// TIA Portal project "Factory_Project_V17" (V17) (continued)
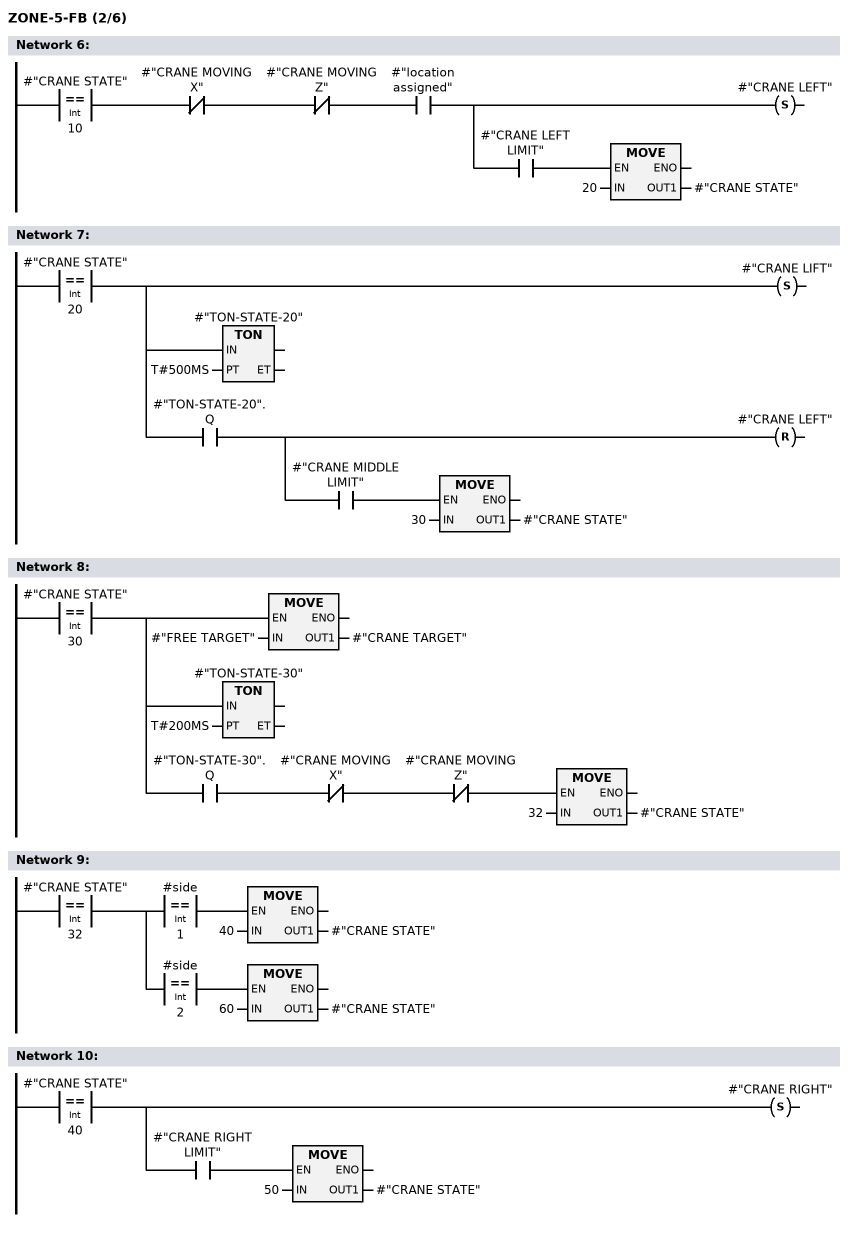
   RUNG wire#powerrail
      { S7_Templates := "SrcType := Int" } EQ_Contact(in1 := #"CRANE STATE", in2 := 10)
      I_Contact( #"CRANE MOVING X" )
      I_Contact( #"CRANE MOVING Z" )
      Contact( #"location assigned" )
      wire#w1
      S_Coil( #"CRANE LEFT" )
   END_RUNG
   RUNG wire#w1
      Contact( #"CRANE LEFT LIMIT" )
      Move(in := 20, out1 => #"CRANE STATE")
   END_RUNG
   // the same network as SCL:
   #_w1 := (#"CRANE STATE" = 10) AND NOT #"CRANE MOVING X" AND NOT #"CRANE MOVING Z" AND #"location assigned";
   IF #_w1 THEN #"CRANE LEFT" := TRUE; END_IF;
   IF #_w1 AND #"CRANE LEFT LIMIT" THEN #"CRANE STATE" := 20; END_IF;
END_REGION

REGION Network 7
   #_w1 := #"CRANE STATE" = 20;
   IF #_w1 THEN #"CRANE LIFT" := TRUE; END_IF;
   #"TON-STATE-20"(IN := #_w1, PT := T#500MS);   // TON
   #_w2 := #_w1 AND #"TON-STATE-20".Q;
   IF #_w2 THEN #"CRANE LEFT" := FALSE; END_IF;
   IF #_w2 AND #"CRANE MIDDLE LIMIT" THEN #"CRANE STATE" := 30; END_IF;
END_REGION

REGION Network 8
   #_w1 := #"CRANE STATE" = 30;
   IF #_w1 THEN #"CRANE TARGET" := #"FREE TARGET"; END_IF;
   #"TON-STATE-30"(IN := #_w1, PT := T#200MS);   // TON
   IF #_w1 AND #"TON-STATE-30".Q AND NOT #"CRANE MOVING X" AND NOT #"CRANE MOVING Z" THEN
       #"CRANE STATE" := 32;
   END_IF;
END_REGION

REGION Network 9
   RUNG wire#powerrail
      { S7_Templates := "SrcType := Int" } EQ_Contact(in1 := #"CRANE STATE", in2 := 32)
      wire#w1
      { S7_Templates := "SrcType := Int" } EQ_Contact(in1 := #side, in2 := 1)
      Move(in := 40, out1 => #"CRANE STATE")
   END_RUNG
   RUNG wire#w1
      { S7_Templates := "SrcType := Int" } EQ_Contact(in1 := #side, in2 := 2)
      Move(in := 60, out1 => #"CRANE STATE")
   END_RUNG
   // the same network as SCL:
   #_w1 := #"CRANE STATE" = 32;
   IF #_w1 AND (#side = 1) THEN #"CRANE STATE" := 40; END_IF;
   IF #_w1 AND (#side = 2) THEN #"CRANE STATE" := 60; END_IF;
END_REGION

REGION Network 10
   RUNG wire#powerrail
      { S7_Templates := "SrcType := Int" } EQ_Contact(in1 := #"CRANE STATE", in2 := 40)
      wire#w1
      S_Coil( #"CRANE RIGHT" )
   END_RUNG
   RUNG wire#w1
      Contact( #"CRANE RIGHT LIMIT" )
      Move(in := 50, out1 => #"CRANE STATE")
   END_RUNG
   // the same network as SCL:
   #_w1 := #"CRANE STATE" = 40;
   IF #_w1 THEN #"CRANE RIGHT" := TRUE; END_IF;
   IF #_w1 AND #"CRANE RIGHT LIMIT" THEN #"CRANE STATE" := 50; END_IF;
END_REGION

REGION Network 11
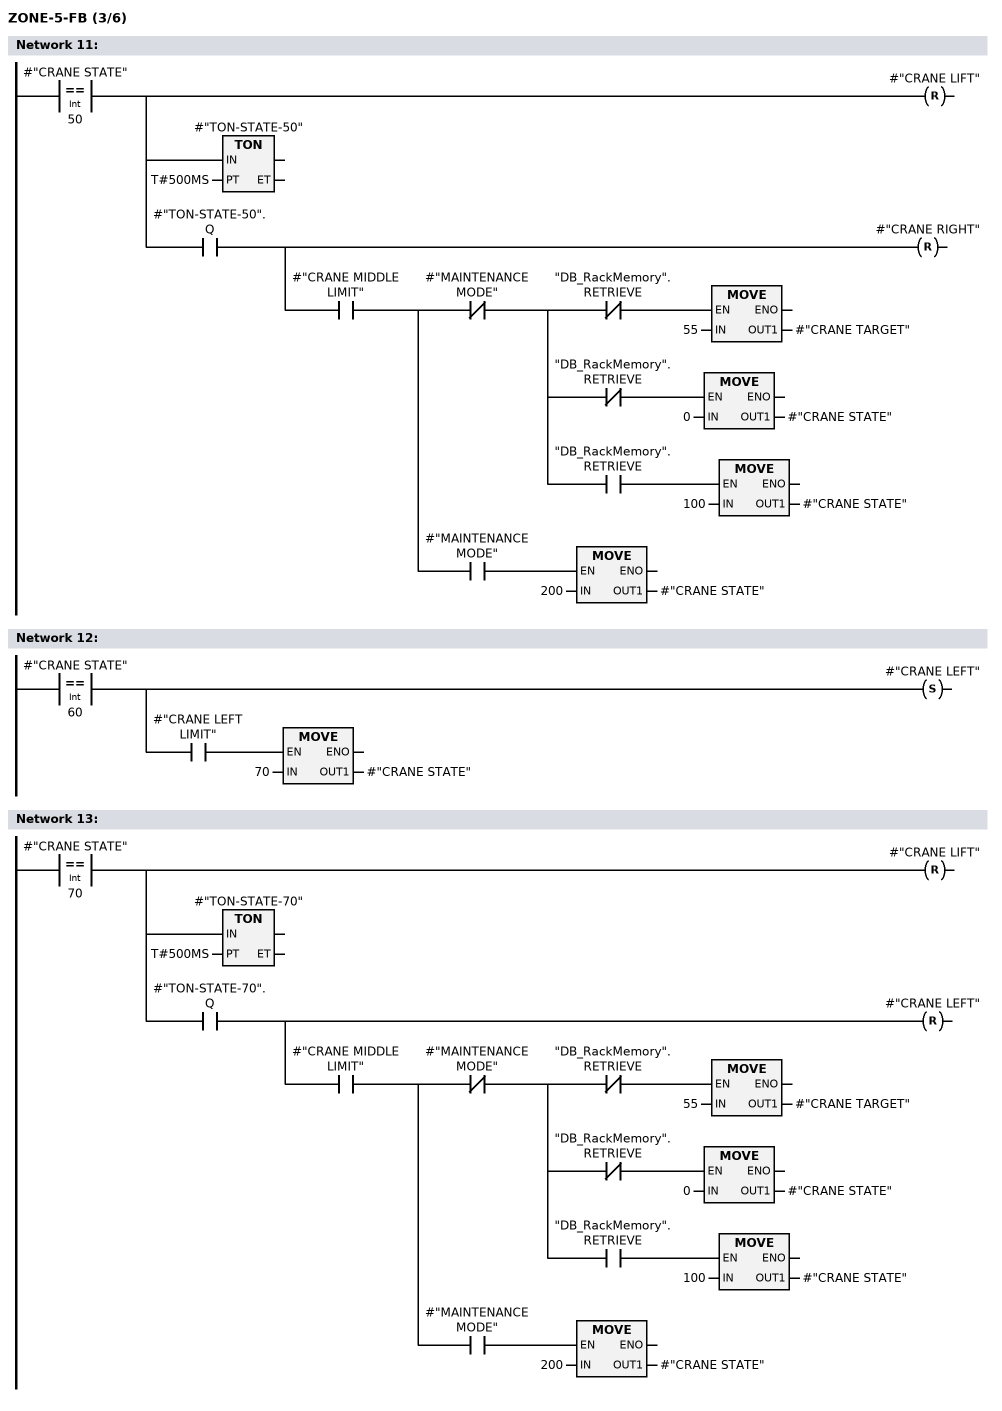
   #_w1 := #"CRANE STATE" = 50;
   IF #_w1 THEN #"CRANE LIFT" := FALSE; END_IF;
   #"TON-STATE-50"(IN := #_w1, PT := T#500MS);   // TON
   #_w2 := #_w1 AND #"TON-STATE-50".Q;
   IF #_w2 THEN #"CRANE RIGHT" := FALSE; END_IF;
   #_w3 := #_w2 AND #"CRANE MIDDLE LIMIT";
   #_w4 := #_w3 AND NOT #"MAINTENANCE MODE";
   IF #_w4 AND NOT "DB_RackMemory".RETRIEVE THEN
       #"CRANE TARGET" := 55;
       #"CRANE STATE" := 0;
   END_IF;
   IF #_w4 AND "DB_RackMemory".RETRIEVE THEN #"CRANE STATE" := 100; END_IF;
   IF #_w3 AND #"MAINTENANCE MODE" THEN #"CRANE STATE" := 200; END_IF;
END_REGION

REGION Network 12
   RUNG wire#powerrail
      { S7_Templates := "SrcType := Int" } EQ_Contact(in1 := #"CRANE STATE", in2 := 60)
      wire#w1
      S_Coil( #"CRANE LEFT" )
   END_RUNG
   RUNG wire#w1
      Contact( #"CRANE LEFT LIMIT" )
      Move(in := 70, out1 => #"CRANE STATE")
   END_RUNG
   // the same network as SCL:
   #_w1 := #"CRANE STATE" = 60;
   IF #_w1 THEN #"CRANE LEFT" := TRUE; END_IF;
   IF #_w1 AND #"CRANE LEFT LIMIT" THEN #"CRANE STATE" := 70; END_IF;
END_REGION

REGION Network 13
   #_w1 := #"CRANE STATE" = 70;
   IF #_w1 THEN #"CRANE LIFT" := FALSE; END_IF;
   #"TON-STATE-70"(IN := #_w1, PT := T#500MS);   // TON
   #_w2 := #_w1 AND #"TON-STATE-70".Q;
   IF #_w2 THEN #"CRANE LEFT" := FALSE; END_IF;
   #_w3 := #_w2 AND #"CRANE MIDDLE LIMIT";
   #_w4 := #_w3 AND NOT #"MAINTENANCE MODE";
   IF #_w4 AND NOT "DB_RackMemory".RETRIEVE THEN
       #"CRANE TARGET" := 55;
       #"CRANE STATE" := 0;
   END_IF;
   IF #_w4 AND "DB_RackMemory".RETRIEVE THEN #"CRANE STATE" := 100; END_IF;
   IF #_w3 AND #"MAINTENANCE MODE" THEN #"CRANE STATE" := 200; END_IF;
END_REGION

REGION Network 14
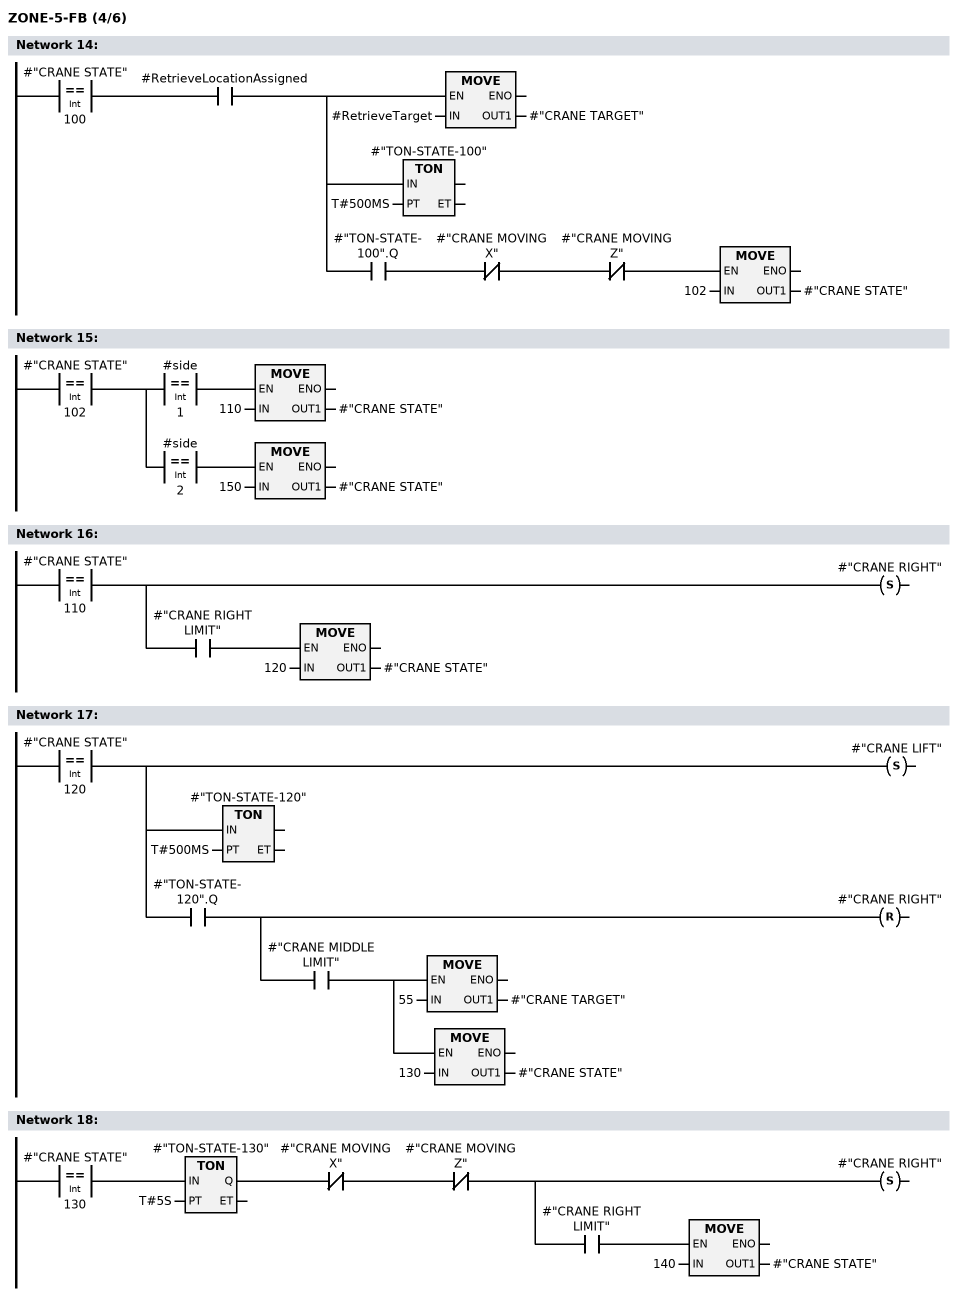
   #_w1 := (#"CRANE STATE" = 100) AND #RetrieveLocationAssigned;
   IF #_w1 THEN #"CRANE TARGET" := #RetrieveTarget; END_IF;
   #"TON-STATE-100"(IN := #_w1, PT := T#500MS);   // TON
   IF #_w1 AND #"TON-STATE-100".Q AND NOT #"CRANE MOVING X" AND NOT #"CRANE MOVING Z" THEN
       #"CRANE STATE" := 102;
   END_IF;
END_REGION

REGION Network 15
   RUNG wire#powerrail
      { S7_Templates := "SrcType := Int" } EQ_Contact(in1 := #"CRANE STATE", in2 := 102)
      wire#w1
      { S7_Templates := "SrcType := Int" } EQ_Contact(in1 := #side, in2 := 1)
      Move(in := 110, out1 => #"CRANE STATE")
   END_RUNG
   RUNG wire#w1
      { S7_Templates := "SrcType := Int" } EQ_Contact(in1 := #side, in2 := 2)
      Move(in := 150, out1 => #"CRANE STATE")
   END_RUNG
   // the same network as SCL:
   #_w1 := #"CRANE STATE" = 102;
   IF #_w1 AND (#side = 1) THEN #"CRANE STATE" := 110; END_IF;
   IF #_w1 AND (#side = 2) THEN #"CRANE STATE" := 150; END_IF;
END_REGION

REGION Network 16
   RUNG wire#powerrail
      { S7_Templates := "SrcType := Int" } EQ_Contact(in1 := #"CRANE STATE", in2 := 110)
      wire#w1
      S_Coil( #"CRANE RIGHT" )
   END_RUNG
   RUNG wire#w1
      Contact( #"CRANE RIGHT LIMIT" )
      Move(in := 120, out1 => #"CRANE STATE")
   END_RUNG
   // the same network as SCL:
   #_w1 := #"CRANE STATE" = 110;
   IF #_w1 THEN #"CRANE RIGHT" := TRUE; END_IF;
   IF #_w1 AND #"CRANE RIGHT LIMIT" THEN #"CRANE STATE" := 120; END_IF;
END_REGION

REGION Network 17
   #_w1 := #"CRANE STATE" = 120;
   IF #_w1 THEN #"CRANE LIFT" := TRUE; END_IF;
   #"TON-STATE-120"(IN := #_w1, PT := T#500MS);   // TON
   #_w2 := #_w1 AND #"TON-STATE-120".Q;
   IF #_w2 THEN #"CRANE RIGHT" := FALSE; END_IF;
   IF #_w2 AND #"CRANE MIDDLE LIMIT" THEN
       #"CRANE TARGET" := 55;
       #"CRANE STATE" := 130;
   END_IF;
END_REGION

REGION Network 18
   #"TON-STATE-130"(IN := #"CRANE STATE" = 130, PT := T#5S);   // TON
   #_w1 := #"TON-STATE-130".Q AND NOT #"CRANE MOVING X" AND NOT #"CRANE MOVING Z";
   IF #_w1 THEN #"CRANE RIGHT" := TRUE; END_IF;
   IF #_w1 AND #"CRANE RIGHT LIMIT" THEN #"CRANE STATE" := 140; END_IF;
END_REGION

REGION Network 19
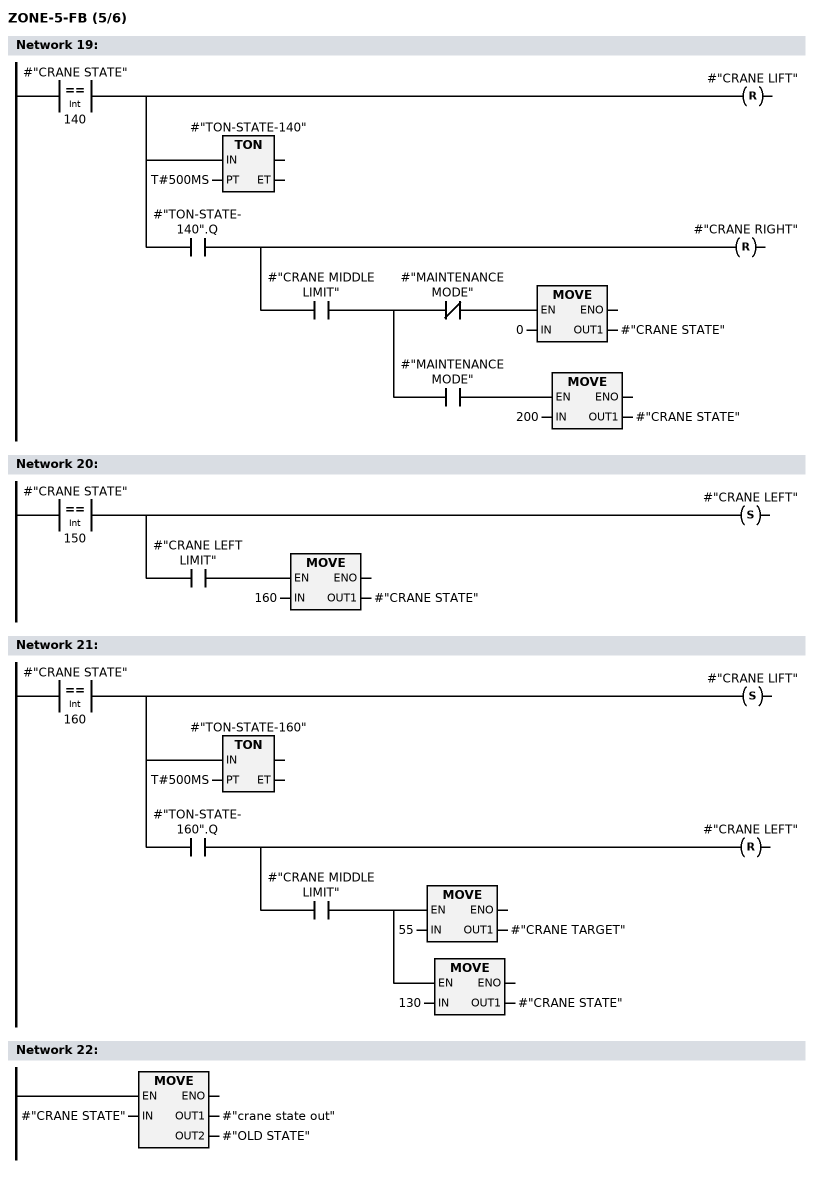
   #_w1 := #"CRANE STATE" = 140;
   IF #_w1 THEN #"CRANE LIFT" := FALSE; END_IF;
   #"TON-STATE-140"(IN := #_w1, PT := T#500MS);   // TON
   #_w2 := #_w1 AND #"TON-STATE-140".Q;
   IF #_w2 THEN #"CRANE RIGHT" := FALSE; END_IF;
   #_w3 := #_w2 AND #"CRANE MIDDLE LIMIT";
   IF #_w3 AND NOT #"MAINTENANCE MODE" THEN #"CRANE STATE" := 0; END_IF;
   IF #_w3 AND #"MAINTENANCE MODE" THEN #"CRANE STATE" := 200; END_IF;
END_REGION

REGION Network 20
   RUNG wire#powerrail
      { S7_Templates := "SrcType := Int" } EQ_Contact(in1 := #"CRANE STATE", in2 := 150)
      wire#w1
      S_Coil( #"CRANE LEFT" )
   END_RUNG
   RUNG wire#w1
      Contact( #"CRANE LEFT LIMIT" )
      Move(in := 160, out1 => #"CRANE STATE")
   END_RUNG
   // the same network as SCL:
   #_w1 := #"CRANE STATE" = 150;
   IF #_w1 THEN #"CRANE LEFT" := TRUE; END_IF;
   IF #_w1 AND #"CRANE LEFT LIMIT" THEN #"CRANE STATE" := 160; END_IF;
END_REGION

REGION Network 21
   #_w1 := #"CRANE STATE" = 160;
   IF #_w1 THEN #"CRANE LIFT" := TRUE; END_IF;
   #"TON-STATE-160"(IN := #_w1, PT := T#500MS);   // TON
   #_w2 := #_w1 AND #"TON-STATE-160".Q;
   IF #_w2 THEN #"CRANE LEFT" := FALSE; END_IF;
   IF #_w2 AND #"CRANE MIDDLE LIMIT" THEN
       #"CRANE TARGET" := 55;
       #"CRANE STATE" := 130;
   END_IF;
END_REGION

REGION Network 22
   RUNG wire#powerrail
      Move(in := #"CRANE STATE", out1 => #"crane state out", out2 => #"OLD STATE")
   END_RUNG
   // the same network as SCL:
   #"crane state out" := #"CRANE STATE";
   #"OLD STATE" := #"CRANE STATE";
END_REGION

REGION Network 23
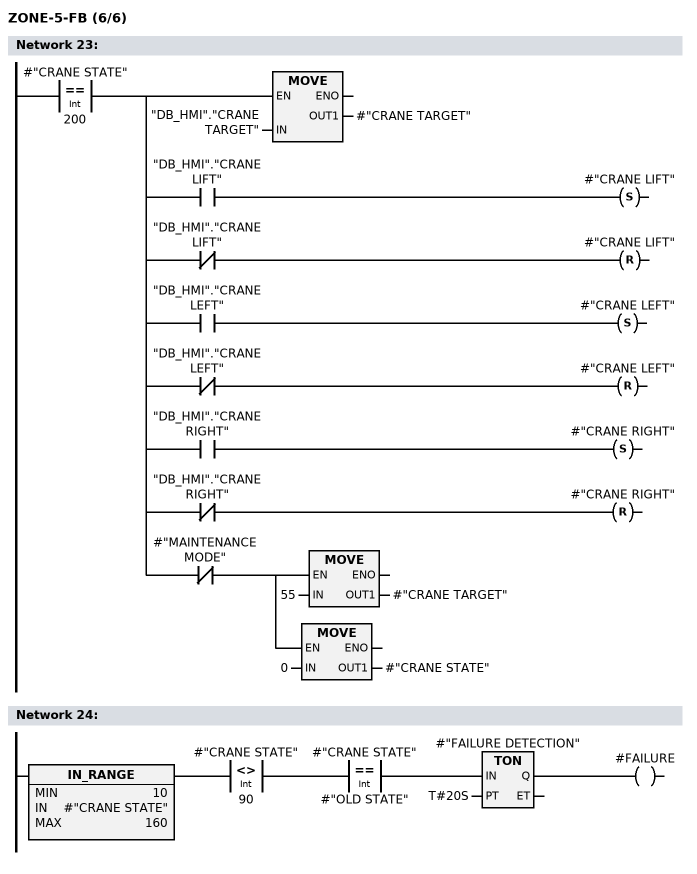
   RUNG wire#powerrail
      { S7_Templates := "SrcType := Int" } EQ_Contact(in1 := #"CRANE STATE", in2 := 200)
      wire#w1
      Move(in := "DB_HMI"."CRANE TARGET", out1 => #"CRANE TARGET")
   END_RUNG
   RUNG wire#w1
      Contact( "DB_HMI"."CRANE LIFT" )
      S_Coil( #"CRANE LIFT" )
   END_RUNG
   RUNG wire#w1
      I_Contact( "DB_HMI"."CRANE LIFT" )
      R_Coil( #"CRANE LIFT" )
   END_RUNG
   RUNG wire#w1
      Contact( "DB_HMI"."CRANE LEFT" )
      S_Coil( #"CRANE LEFT" )
   END_RUNG
   RUNG wire#w1
      I_Contact( "DB_HMI"."CRANE LEFT" )
      R_Coil( #"CRANE LEFT" )
   END_RUNG
   RUNG wire#w1
      Contact( "DB_HMI"."CRANE RIGHT" )
      S_Coil( #"CRANE RIGHT" )
   END_RUNG
   RUNG wire#w1
      I_Contact( "DB_HMI"."CRANE RIGHT" )
      R_Coil( #"CRANE RIGHT" )
   END_RUNG
   RUNG wire#w1
      I_Contact( #"MAINTENANCE MODE" )
      wire#w2
      Move(in := 55, out1 => #"CRANE TARGET")
   END_RUNG
   RUNG wire#w2
      Move(in := 0, out1 => #"CRANE STATE")
   END_RUNG
   // the same network as SCL:
   #_w1 := #"CRANE STATE" = 200;
   IF #_w1 THEN #"CRANE TARGET" := "DB_HMI"."CRANE TARGET"; END_IF;
   IF #_w1 AND "DB_HMI"."CRANE LIFT" THEN #"CRANE LIFT" := TRUE; END_IF;
   IF #_w1 AND NOT "DB_HMI"."CRANE LIFT" THEN #"CRANE LIFT" := FALSE; END_IF;
   IF #_w1 AND "DB_HMI"."CRANE LEFT" THEN #"CRANE LEFT" := TRUE; END_IF;
   IF #_w1 AND NOT "DB_HMI"."CRANE LEFT" THEN #"CRANE LEFT" := FALSE; END_IF;
   IF #_w1 AND "DB_HMI"."CRANE RIGHT" THEN #"CRANE RIGHT" := TRUE; END_IF;
   IF #_w1 AND NOT "DB_HMI"."CRANE RIGHT" THEN #"CRANE RIGHT" := FALSE; END_IF;
   IF #_w1 AND NOT #"MAINTENANCE MODE" THEN
       #"CRANE TARGET" := 55;
       #"CRANE STATE" := 0;
   END_IF;
END_REGION

REGION Network 24
   #"FAILURE DETECTION"(IN := (10 <= #"CRANE STATE") AND (#"CRANE STATE" <= 160) AND (#"CRANE STATE" <> 90) AND (#"CRANE STATE" = #"OLD STATE"),   // TON
                        PT := T#20S);
   #FAILURE := #"FAILURE DETECTION".Q;
END_REGION
END_FUNCTION_BLOCK

// folder: ZONE-5-BLOCKS/ZONE 5 SUB BLOCKS

FUNCTION_BLOCK "RACK MANAGMENT"   // FB20, SCL
{ S7_Optimized_Access := 'TRUE' }
VERSION : 0.1
   VAR_INPUT
      "crane state" : Int;
      RetireveQuantity : Int;
      cancel : Bool;
      "RESET MEMORY" : Bool;
   END_VAR
   VAR_OUTPUT
      target : Int;
      side : Int;
      warehouse_full : Bool;
      location_assigned : Bool;
      RetrieveTarget : Int;
      RetrieveSide : Int;
      RetrieveLocationAssigned : Bool;
      "FREE SPACES" : Int;
   END_VAR
   VAR
      i : Int;
      found : Bool;
      j : Int;
      RetireveFound : Bool;
      RETRIEVE_R_TRIG_Instance : R_TRIG;
      "RETRIEVE P TRIG" : Bool;
   END_VAR
BEGIN
   #RETRIEVE_R_TRIG_Instance(CLK:="DB_RackMemory".RETRIEVE,
                             Q=>#"RETRIEVE P TRIG");

   IF NOT #warehouse_full THEN
       IF #"crane state" = 10 AND NOT #location_assigned THEN
           #found := FALSE;
           FOR #i := 1 TO 108 DO
               IF NOT "DB_RackMemory".Rack[#i].occupied THEN
                   #target := #i;
                   #side := "DB_RackMemory".Rack[#i].side;
                   #found := TRUE;
                   EXIT;
               END_IF;
           END_FOR;

           IF NOT #found THEN
               #warehouse_full := TRUE;
           ELSE
               #location_assigned := TRUE;
           END_IF;

       END_IF;
       IF #"crane state" = 50 AND #location_assigned THEN
           "DB_RackMemory".Rack[#i].occupied := TRUE;

           #location_assigned := FALSE;
       END_IF;
   END_IF;
   IF #"RETRIEVE P TRIG" THEN
       "DB_RackMemory"."REQUIRED QUANTITY" := "DB_RackMemory"."QUANTITY TO RETRIEVE";
   END_IF;
   IF "DB_RackMemory".RETRIEVE AND "DB_RackMemory"."QUANTITY TO RETRIEVE" > 0 THEN
       IF #"crane state" = 100 AND NOT #RetrieveLocationAssigned THEN
           #RetireveFound := FALSE;
           FOR #i := 1 TO 108 DO
               IF "DB_RackMemory".Rack[#i].occupied THEN
                   #RetrieveTarget := #i;
                   #RetrieveSide := "DB_RackMemory".Rack[#i].side;
                   #RetireveFound := TRUE;
                   EXIT;
               END_IF;
           END_FOR;

           #RetrieveLocationAssigned := TRUE;
       END_IF;

       IF #"crane state" = 140 AND #RetrieveLocationAssigned THEN
           "DB_RackMemory".Rack[#i].occupied := FALSE;
           "DB_RackMemory".SpacesOccupied := "DB_RackMemory".SpacesOccupied - 1;
           "DB_RackMemory"."QUANTITY TO RETRIEVE" := "DB_RackMemory"."QUANTITY TO RETRIEVE" - 1;
           "DB_RackMemory"."TOTAL DLIEVERED" := "DB_RackMemory"."TOTAL DLIEVERED" + 1;

           IF "DB_RackMemory"."QUANTITY TO RETRIEVE" = 0 THEN
               "DB_RackMemory".RETRIEVE := FALSE;
               "DB_RackMemory"."TOTAL ORDERS" := "DB_RackMemory"."TOTAL ORDERS" + 1;
               "DB_RackMemory"."REQUIRED QUANTITY" := 0;
           END_IF;
           #RetrieveLocationAssigned := FALSE;
           IF #warehouse_full THEN
               #warehouse_full := FALSE;
           END_IF;
           IF #cancel THEN
               "DB_RackMemory".RETRIEVE := FALSE;
               "DB_RackMemory"."QUANTITY TO RETRIEVE" := 0;
               "DB_HMI"."CANCEL ORDER" := FALSE;
           END_IF;
       END_IF;
   END_IF;
   #"FREE SPACES" := 108 - "DB_RackMemory".SpacesOccupied;
   IF "DB_RackMemory".RETRIEVE AND "DB_RackMemory"."QUANTITY TO RETRIEVE" = 0 THEN
       "DB_RackMemory".RETRIEVE := FALSE;
   END_IF;
   IF #"RESET MEMORY" THEN
       "DB_RackMemory"."QUANTITY TO RETRIEVE" := 0;
       "DB_RackMemory"."REQUIRED QUANTITY" := 0;
       "DB_RackMemory".SpacesOccupied := 0;
       "DB_RackMemory"."TOTAL ORDERS" := 0;
       "DB_RackMemory"."TOTAL DLIEVERED" := 0;
       "DB_RackMemory".RETRIEVE := FALSE;
       FOR #i := 1 TO 108 DO
           "DB_RackMemory".Rack[#i].occupied := FALSE;
       END_FOR;
       "DB_RackMemory".ReckMemoryReset := FALSE;
   END_IF;
END_FUNCTION_BLOCK

// folder: ZONE_1_BLOCKS

FUNCTION_BLOCK "Zone_1_FB"   // FB1, LAD
{ S7_Optimized_Access := 'TRUE' }
VERSION : 0.1
   VAR_INPUT
      SystemEnabled : Bool;
      stop : Bool;
      EMERGENCY : Bool;
      EntrySensor : Bool;
      AtScaleSensor : Bool;
      VisionSensor : Bool;
      ScaleValue : Real;
      reset : Bool;
      "machine A entry" : Bool;
      "machine B entry" : Bool;
   END_VAR
   VAR_OUTPUT
      Emitter : Bool;
      "sorter left" : Bool;
      "sorter right" : Bool;
      feed_conv : Bool;
      Z1L1 : Bool;
      Z1L2 : Bool;
      Z1L3 : Bool;
      Z1L4 : Bool;
      Z1L5 : Bool;
      Z1L6 : Bool;
      Z1L7 : Bool;
      Z1L8 : Bool;
      Z1R1 : Bool;
      Z1R2 : Bool;
      Z1R3 : Bool;
      Z1R4 : Bool;
      Z1R5 : Bool;
      Z1R6 : Bool;
      scale_conv : Bool;
      sorter_wheels : Bool;
      Zone1_state : Int;
   END_VAR
   VAR
      STATE : Int;
      DecisionPulse : Bool;
      "l/r" : Int;
      toggle_Instance : "toggle";
      decision : Int;
      currentState : Int;
      stopped : Bool;
      Z1_Sorter_Decision_fb_Instance : "Z1_Sorter_Decision_fb";
      Z1_Conv_Activation_FB_Instance : "Z1_Conv_Activation_FB";
      Z1_Reset_Program_Instance : "Z1_Reset_Program";
      reset_timer : Bool;
      reset_timer_0 : TON_TIME;
   END_VAR
   VAR RETAIN
      IEC_Counter_0_Instance : CTU_INT;
      "CTU-IN-PRODUCTION" : CTU_INT;
      "L/R IS ZERO" : Bool;
      "L/R IS ONE" : Bool;
   END_VAR
   VAR
      "CTU-PRODUCTION-RESET" : Bool;
      "PRODUCTION LIMIT_Instance" : "PRODUCTION LIMIT";
      "LIMIT REACHED" : Bool;
   END_VAR
   VAR_TEMP
      reset_complete : Bool;
      Temp_1 : Bool;
   END_VAR
   VAR_TEMP   // added for the SCL form of the ladder/FBD networks
      _w1 : Bool;
      _w2 : Bool;
      _w3 : Bool;
      _w4 : Bool;
   END_VAR
BEGIN

REGION Network 1
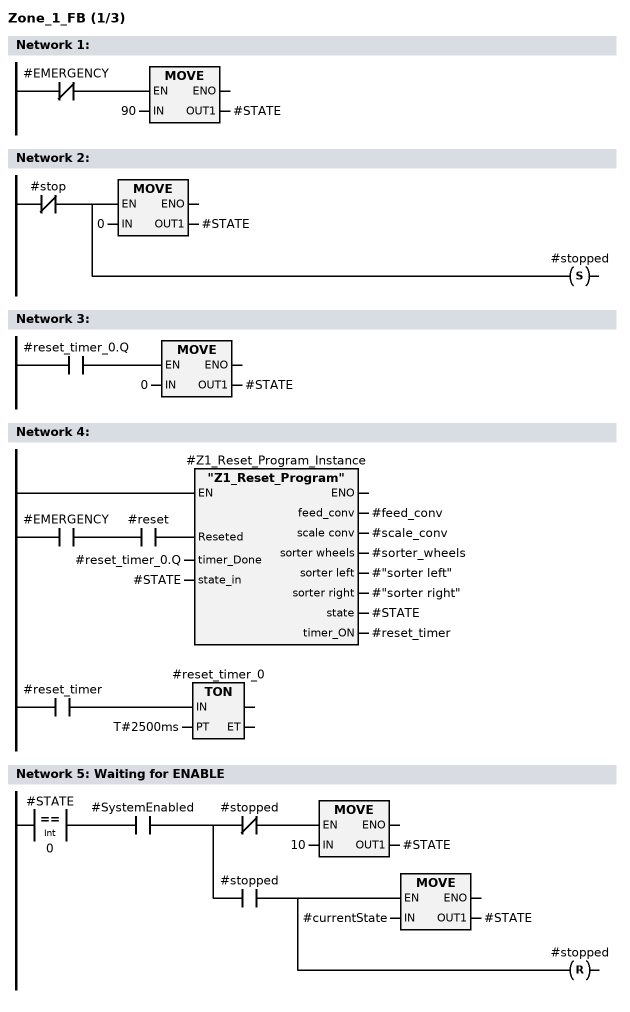
   RUNG wire#powerrail
      I_Contact( #EMERGENCY )
      Move(in := 90, out1 => #STATE)
   END_RUNG
   // the same network as SCL:
   IF NOT #EMERGENCY THEN #STATE := 90; END_IF;
END_REGION

REGION Network 2
   RUNG wire#powerrail
      I_Contact( #stop )
      wire#w1
      Move(in := 0, out1 => #STATE)
   END_RUNG
   RUNG wire#w1
      S_Coil( #stopped )
   END_RUNG
   // the same network as SCL:
   IF NOT #stop THEN
       #STATE := 0;
       #stopped := TRUE;
   END_IF;
END_REGION

REGION Network 3
   RUNG wire#powerrail
      Contact( #reset_timer_0.Q )
      Move(in := 0, out1 => #STATE)
   END_RUNG
   // the same network as SCL:
   IF #reset_timer_0.Q THEN #STATE := 0; END_IF;
END_REGION

REGION Network 4
   #Z1_Reset_Program_Instance(Reseted := #EMERGENCY AND #reset,   // "Z1_Reset_Program"
                           timer_Done := #reset_timer_0.Q,
                           state_in := #STATE,
                           feed_conv => #feed_conv,
                           "scale conv" => #scale_conv,
                           "sorter wheels" => #sorter_wheels,
                           "sorter left" => #"sorter left",
                           "sorter right" => #"sorter right",
                           state => #STATE,
                           timer_ON => #reset_timer);
   #reset_timer_0(IN := #reset_timer, PT := T#2500ms);   // TON
END_REGION

REGION Network 5: Waiting for ENABLE
   RUNG wire#powerrail
      { S7_Templates := "SrcType := Int" } EQ_Contact(in1 := #STATE, in2 := 0)
      Contact( #SystemEnabled )
      wire#w1
      I_Contact( #stopped )
      Move(in := 10, out1 => #STATE)
   END_RUNG
   RUNG wire#w1
      Contact( #stopped )
      wire#w2
      Move(in := #currentState, out1 => #STATE)
   END_RUNG
   RUNG wire#w2
      R_Coil( #stopped )
   END_RUNG
   // the same network as SCL:
   #_w1 := (#STATE = 0) AND #SystemEnabled;
   IF #_w1 AND NOT #stopped THEN #STATE := 10; END_IF;
   IF #_w1 AND #stopped THEN
       #STATE := #currentState;
       #stopped := FALSE;
   END_IF;
END_REGION

REGION Network 6
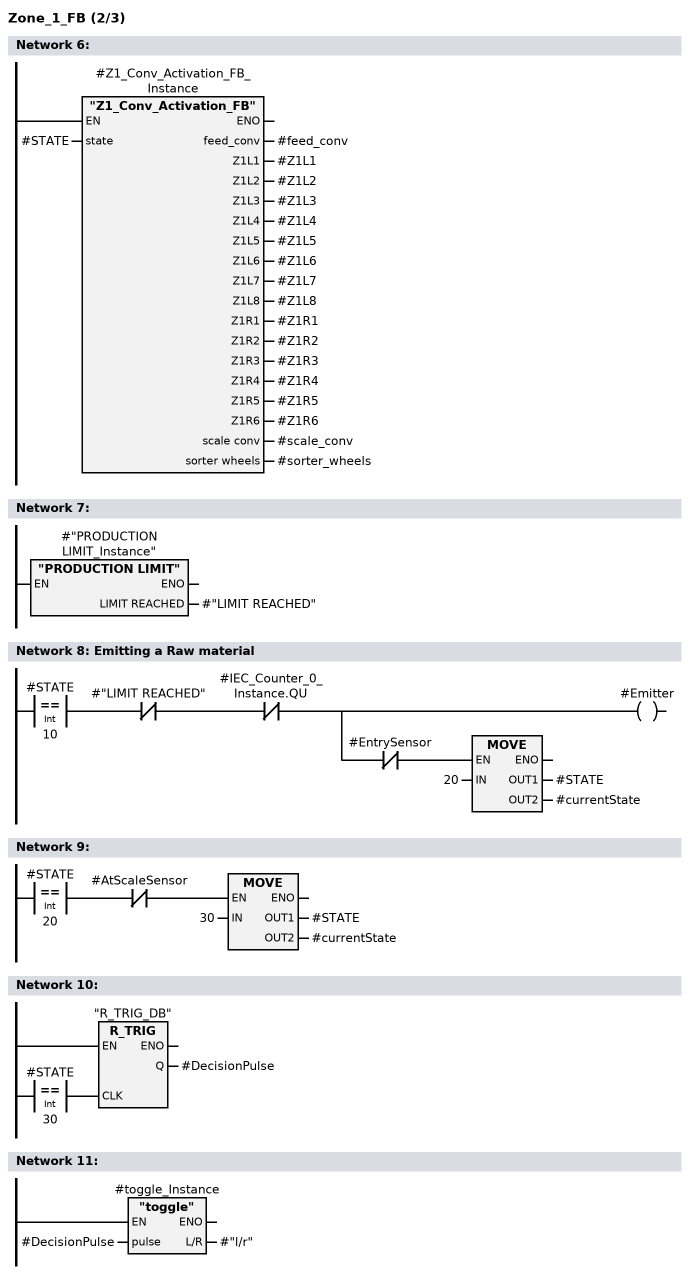
   RUNG wire#powerrail
      #Z1_Conv_Activation_FB_Instance(state := #STATE, feed_conv => #feed_conv, Z1L1 => #Z1L1, Z1L2 => #Z1L2, Z1L3 => #Z1L3, Z1L4 => #Z1L4, Z1L5 => #Z1L5, Z1L6 => #Z1L6, Z1L7 => #Z1L7, Z1L8 => #Z1L8, Z1R1 => #Z1R1, Z1R2 => #Z1R2, Z1R3 => #Z1R3, Z1R4 => #Z1R4, Z1R5 => #Z1R5, Z1R6 => #Z1R6, "scale conv" => #scale_conv, "sorter wheels" => #sorter_wheels)
   END_RUNG
   // the same network as SCL:
   #Z1_Conv_Activation_FB_Instance(state := #STATE,   // "Z1_Conv_Activation_FB"
                           feed_conv => #feed_conv,
                           Z1L1 => #Z1L1,
                           Z1L2 => #Z1L2,
                           Z1L3 => #Z1L3,
                           Z1L4 => #Z1L4,
                           Z1L5 => #Z1L5,
                           Z1L6 => #Z1L6,
                           Z1L7 => #Z1L7,
                           Z1L8 => #Z1L8,
                           Z1R1 => #Z1R1,
                           Z1R2 => #Z1R2,
                           Z1R3 => #Z1R3,
                           Z1R4 => #Z1R4,
                           Z1R5 => #Z1R5,
                           Z1R6 => #Z1R6,
                           "scale conv" => #scale_conv,
                           "sorter wheels" => #sorter_wheels);
END_REGION

REGION Network 7
   RUNG wire#powerrail
      #"PRODUCTION LIMIT_Instance"("LIMIT REACHED" => #"LIMIT REACHED")
   END_RUNG
   // the same network as SCL:
   #"PRODUCTION LIMIT_Instance"("LIMIT REACHED" => #"LIMIT REACHED");   // "PRODUCTION LIMIT"
END_REGION

REGION Network 8: Emitting a Raw material
   RUNG wire#powerrail
      { S7_Templates := "SrcType := Int" } EQ_Contact(in1 := #STATE, in2 := 10)
      I_Contact( #"LIMIT REACHED" )
      I_Contact( #IEC_Counter_0_Instance.QU )
      wire#w1
      Coil( #Emitter )
   END_RUNG
   RUNG wire#w1
      I_Contact( #EntrySensor )
      Move(in := 20, out1 => #STATE, out2 => #currentState)
   END_RUNG
   // the same network as SCL:
   #Emitter := (#STATE = 10) AND NOT #"LIMIT REACHED" AND NOT #IEC_Counter_0_Instance.QU;
   IF #Emitter AND NOT #EntrySensor THEN
       #STATE := 20;
       #currentState := 20;
   END_IF;
END_REGION

REGION Network 9
   RUNG wire#powerrail
      { S7_Templates := "SrcType := Int" } EQ_Contact(in1 := #STATE, in2 := 20)
      I_Contact( #AtScaleSensor )
      Move(in := 30, out1 => #STATE, out2 => #currentState)
   END_RUNG
   // the same network as SCL:
   IF (#STATE = 20) AND NOT #AtScaleSensor THEN
       #STATE := 30;
       #currentState := 30;
   END_IF;
END_REGION

REGION Network 10
   "R_TRIG_DB"(CLK := #STATE = 30, Q => #DecisionPulse);   // R_TRIG
END_REGION

REGION Network 11
   RUNG wire#powerrail
      #toggle_Instance(pulse := #DecisionPulse, "L/R" => #"l/r")
   END_RUNG
   // the same network as SCL:
   #toggle_Instance(pulse := #DecisionPulse, "L/R" => #"l/r");   // "toggle"
END_REGION

REGION Network 12
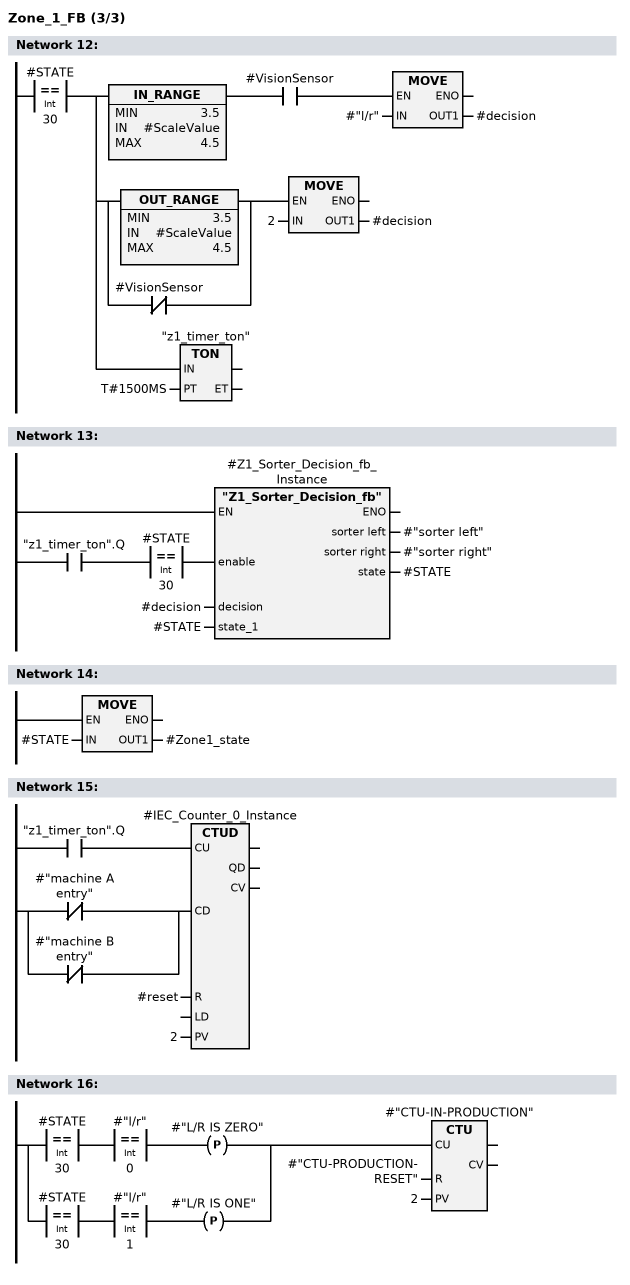
   #_w1 := #STATE = 30;
   IF #_w1 AND (3.5 <= #ScaleValue) AND (#ScaleValue <= 4.5) AND #VisionSensor THEN
       #decision := #"l/r";
   END_IF;
   IF #_w1 AND ((#ScaleValue < 3.5) OR (#ScaleValue > 4.5) OR NOT #VisionSensor) THEN #decision := 2; END_IF;
   "z1_timer_ton".TON(IN := #_w1, PT := T#1500MS);
END_REGION

REGION Network 13
   RUNG wire#powerrail
      #Z1_Sorter_Decision_fb_Instance(enable := wire#w1, decision := #decision, state_1 := #STATE, "sorter left" => #"sorter left", "sorter right" => #"sorter right", state => #STATE)
   END_RUNG
   RUNG wire#powerrail
      Contact( "z1_timer_ton".Q )
      { S7_Templates := "SrcType := Int" } EQ_Contact(in1 := #STATE, in2 := 30)
   END_RUNG wire#w1
   // the same network as SCL:
   #Z1_Sorter_Decision_fb_Instance(enable := "z1_timer_ton".Q AND (#STATE = 30),   // "Z1_Sorter_Decision_fb"
                           decision := #decision,
                           state_1 := #STATE,
                           "sorter left" => #"sorter left",
                           "sorter right" => #"sorter right",
                           state => #STATE);
END_REGION

REGION Network 14
   RUNG wire#powerrail
      Move(in := #STATE, out1 => #Zone1_state)
   END_RUNG
   // the same network as SCL:
   #Zone1_state := #STATE;
END_REGION

REGION Network 15
   #IEC_Counter_0_Instance(CU := "z1_timer_ton".Q,   // CTUD
                           CD := NOT #"machine A entry" OR NOT #"machine B entry",
                           R := #reset,
                           PV := 2);
END_REGION

REGION Network 16
   #_w1 := (#STATE = 30) AND (#"l/r" = 0);
   #_w2 := #_w1 AND NOT #"L/R IS ZERO";   // rising edge
   #"L/R IS ZERO" := #_w1;
   #_w3 := (#STATE = 30) AND (#"l/r" = 1);
   #_w4 := #_w3 AND NOT #"L/R IS ONE";   // rising edge
   #"L/R IS ONE" := #_w3;
   #"CTU-IN-PRODUCTION"(CU := #_w2 OR #_w4, R := #"CTU-PRODUCTION-RESET", PV := 2);   // CTU
END_REGION

REGION Network 17 (SCL)
   IF #"CTU-IN-PRODUCTION".QU THEN
       "DB_RackMemory".In_Production := "DB_RackMemory".In_Production + 1;
       #"CTU-PRODUCTION-RESET" := TRUE;
   ELSE
       #"CTU-PRODUCTION-RESET" := FALSE;
   END_IF;
END_REGION

REGION Network 18 (SCL)
   IF "DB_RackMemory".InProductionReset THEN
       "DB_RackMemory".In_Production := 0;
       "DB_RackMemory".InProductionReset := FALSE;
   END_IF;
END_REGION
END_FUNCTION_BLOCK

// folder: ZONE_1_BLOCKS/ZONE 1 SUB BLOCKS

FUNCTION_BLOCK "toggle"   // FB2, SCL
{ S7_Optimized_Access := 'TRUE' }
VERSION : 0.1
   VAR_INPUT
      pulse : Bool;
   END_VAR
   VAR_OUTPUT
      "L/R" : Int;
   END_VAR
   VAR
      to_toggle : Bool;
   END_VAR
BEGIN
   IF #pulse THEN
       // Statement section IF
       #to_toggle:= NOT #to_toggle;
       IF #to_toggle THEN
           #"L/R" := 1;
       END_IF;
       IF NOT #to_toggle THEN
           #"L/R" := 0;
       END_IF;
   END_IF;
END_FUNCTION_BLOCK

FUNCTION_BLOCK "Z1_Sorter_Decision_fb"   // FB3, SCL
{ S7_Optimized_Access := 'TRUE' }
VERSION : 0.1
   VAR_INPUT
      enable : Bool;
      decision : Int;
      state_1 : Int;
   END_VAR
   VAR_OUTPUT
      "sorter left" : Bool;
      "sorter right" : Bool;
      state : Int;
   END_VAR
BEGIN
   IF #enable THEN
       // Statement section IF
       CASE #decision OF
           0:  // Statement section case 1
               #"sorter left" := 1;
               #"sorter right" := 0;
               #state := 10;
           1:  // Statement section case 2 to 4
               #"sorter left":= 0;
               #"sorter right" := 1;
               #state := 10;
           2:
               #"sorter left" := 0;
               #"sorter right" := 0;
               #state := 10;
           ELSE  // Statement section ELSE
               #"sorter left" := 0;
               #"sorter right" := 0;
               #state := 100;
       END_CASE;
   ELSIF #state_1 = 100 OR #state_1=90  THEN
       #state := #state_1;
       #"sorter left" := 0;
       #"sorter right" := 0;
   ELSIF #state_1 = 0 THEN
       #state := #state_1;
       #"sorter left" := 0;
       #"sorter right" := 0;
   ELSE
       #state := #state_1;
   END_IF;
END_FUNCTION_BLOCK

FUNCTION_BLOCK "Z1_Conv_Activation_FB"   // FB4, SCL
{ S7_Optimized_Access := 'TRUE' }
VERSION : 0.1
   VAR_INPUT
      state : Int;
   END_VAR
   VAR_OUTPUT
      feed_conv : Bool;
      Z1L1 : Bool;
      Z1L2 : Bool;
      Z1L3 : Bool;
      Z1L4 : Bool;
      Z1L5 : Bool;
      Z1L6 : Bool;
      Z1L7 : Bool;
      Z1L8 : Bool;
      Z1R1 : Bool;
      Z1R2 : Bool;
      Z1R3 : Bool;
      Z1R4 : Bool;
      Z1R5 : Bool;
      Z1R6 : Bool;
      "scale conv" : Bool;
      "sorter wheels" : Bool;
   END_VAR
BEGIN
   IF #state = 10 OR #state = 20 THEN
       // Statement section IF
       #feed_conv := 1;
       #Z1L1 := 1;
       #Z1L2 := 1;
       #Z1L3 := 1;
       #Z1L4 := 1;
       #Z1L5 := 1;
       #Z1L6 := 1;
       #Z1L7 := 1;
       #Z1L8 := 1;
       #Z1R1 := 1;
       #Z1R2 := 1;
       #Z1R3 := 1;
       #Z1R4 := 1;
       #Z1R5 := 1;
       #Z1R6 := 1;
       #"scale conv" := 1;
       #"sorter wheels" := 1;
   END_IF;
   IF #state = 30 THEN
       #feed_conv := 1;
       #Z1L1 := 1;
       #Z1L2 := 1;
       #Z1L3 := 1;
       #Z1L4 := 1;
       #Z1L5 := 1;
       #Z1L6 := 1;
       #Z1L7 := 1;
       #Z1L8 := 1;
       #Z1R1 := 1;
       #Z1R2 := 1;
       #Z1R3 := 1;
       #Z1R4 := 1;
       #Z1R5 := 1;
       #Z1R6 := 1;
       #"sorter wheels" := 1;
       #"scale conv" := 0;
   END_IF;
   IF #state = 0 OR #state=90 THEN
           #feed_conv := 0;
           #Z1L1 := 0;
           #Z1L2 := 0;
           #Z1L3 := 0;
           #Z1L4 := 0;
           #Z1L5 := 0;
           #Z1L6 := 0;
           #Z1L7 := 0;
           #Z1L8 := 0;
           #Z1R1 := 0;
           #Z1R2 := 0;
           #Z1R3 := 0;
           #Z1R4 := 0;
           #Z1R5 := 0;
           #Z1R6 := 0;
           #"sorter wheels" := 0;
           #"scale conv" := 0;
   END_IF;
   IF #state = 100 THEN

       #"scale conv" := 1;
   END_IF;
END_FUNCTION_BLOCK

FUNCTION_BLOCK "Z1_Reset_Program"   // FB5, SCL
{ S7_Optimized_Access := 'TRUE' }
VERSION : 0.1
   VAR_INPUT
      Reseted : Bool;
      timer_Done : Bool;
      state_in : Int;
   END_VAR
   VAR_OUTPUT
      feed_conv : Bool;
      "scale conv" : Bool;
      "sorter wheels" : Bool;
      "sorter left" : Bool;
      "sorter right" : Bool;
      state : Int;
      timer_ON : Bool;
   END_VAR
BEGIN
   IF #Reseted THEN
       // Statement section IF
       #feed_conv := 1;
       #"scale conv" := 1;
       #"sorter wheels" := 1;
       #"sorter left" := 1;
       #"sorter right" := 1;
       #timer_ON := 1;
       #state := 100;
   ELSE
       #state := #state_in;
   END_IF;
   IF #timer_Done THEN
       #feed_conv := 0;
       #"scale conv" := 0;
       #"sorter wheels" := 0;
       #"sorter left" := 0;
       #"sorter right" := 0;
       #timer_ON := 0;

   END_IF;
END_FUNCTION_BLOCK

FUNCTION_BLOCK "PRODUCTION LIMIT"   // FB21, SCL
{ S7_Optimized_Access := 'TRUE' }
VERSION : 0.1
   VAR_OUTPUT
      "LIMIT REACHED" : Bool;
   END_VAR
BEGIN
   IF (("DB_RackMemory".In_Production / 2) + "DB_RackMemory".SpacesOccupied) = 108 THEN
       #"LIMIT REACHED" := TRUE;
   END_IF;
   IF #"LIMIT REACHED" AND (("DB_RackMemory".In_Production / 2) + "DB_RackMemory".SpacesOccupied) <= 102 THEN
       #"LIMIT REACHED" := FALSE;
   END_IF;
END_FUNCTION_BLOCK

// folder: ZONE_4_BLOCKS

FUNCTION_BLOCK "ZONE 4 FB"   // FB16, LAD
{ S7_Optimized_Access := 'TRUE' }
VERSION : 0.1
   VAR_INPUT
      "PALLETIZER ELEVATOR BACK LIMIT" : Bool;
      "PALLETIZER ELEVATOR FRONT LIMIT" : Bool;
      "ELEVATOR MOVING" : Bool;
      "PLATE LIMIT" : Bool;
      "PUSHER LIMIT" : Bool;
      "PALLETIZER ENTRY" : Bool;
      RESET : Bool;
      EMERGENCY : Bool;
   END_VAR
   VAR_OUTPUT
      TURN : Bool;
      PUSH : Bool;
      CLAMP : Bool;
      "OPEN PLATE" : Bool;
      "BELT +" : Bool;
      "CHAIN +" : Bool;
      "ELEVATOR +" : Bool;
      "ELEVATOR -" : Bool;
      "ELEVATOR TO LIMIT" : Bool;
      "PALLETIZER EMITTER" : Bool;
      FAILURE : Bool;
   END_VAR
   VAR
      "PALLETIZER STATE" : Int;
      "ENTRY SENSOR TRIGGER BIT" : Bool;
   END_VAR
   VAR RETAIN
      "CTUD-0" : CTUD_INT;
      "CTUD-1" : CTUD_INT;
   END_VAR
   VAR
      "TON-STATE-30" : TON_TIME;
      "TON-STATE-40" : TON_TIME;
      "LOWER PART READY" : Bool;
      "UPPER READY" : Bool;
      "ZONE 4 LOWER PART LOGIC_Instance" : "ZONE 4 LOWER PART LOGIC";
      "TON-STATE-10-A" : TON_TIME;
      "TON-STATE-10-B" : TON_TIME;
      "TON-STATE-12" : TON_TIME;
      "TON-STATE-0" : TON_TIME;
      "TON-STATE-20" : TON_TIME;
      "TON-STATE-40-B" : TON_TIME;
      "PRODUCTS UPDATE" : Bool;
      "OLD STATE" : Int;
      "FAILURE DETECTION" : TON_TIME;
      "UPPER FAIL" : Bool;
      "LOWER FAIL" : Bool;
   END_VAR
   VAR_TEMP   // added for the SCL form of the ladder/FBD networks
      _w1 : Bool;
      _w2 : Bool;
   END_VAR
BEGIN

REGION Network 1